// TIA Portal project "1215C_BREAKOUT_BOARD_IO-LINK_TOWERLIGHT" (V19) (continued)
REGION Network 1: ================= PORT_X1 =================
END_REGION

REGION Network 2: Reserved
END_REGION

REGION Network 3: ================= PORT_X2 =================
END_REGION

REGION Network 4: Banner Tower Light
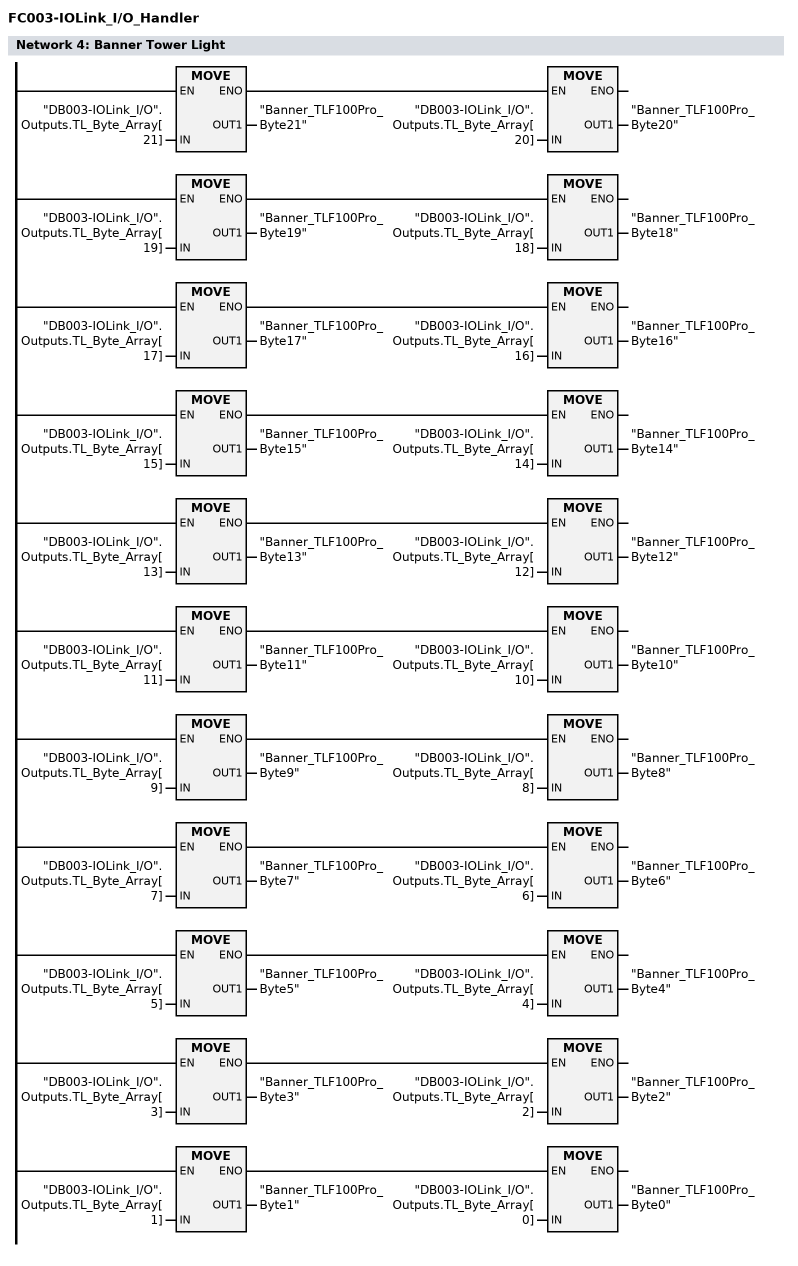
   RUNG wire#powerrail
      Move(in := "DB003-IOLink_I/O".Outputs.TL_Byte_Array[21], out1 => "Banner_TLF100Pro_Byte21")
      Move(in := "DB003-IOLink_I/O".Outputs.TL_Byte_Array[20], out1 => "Banner_TLF100Pro_Byte20")
   END_RUNG
   RUNG wire#powerrail
      Move(in := "DB003-IOLink_I/O".Outputs.TL_Byte_Array[19], out1 => "Banner_TLF100Pro_Byte19")
      Move(in := "DB003-IOLink_I/O".Outputs.TL_Byte_Array[18], out1 => "Banner_TLF100Pro_Byte18")
   END_RUNG
   RUNG wire#powerrail
      Move(in := "DB003-IOLink_I/O".Outputs.TL_Byte_Array[17], out1 => "Banner_TLF100Pro_Byte17")
      Move(in := "DB003-IOLink_I/O".Outputs.TL_Byte_Array[16], out1 => "Banner_TLF100Pro_Byte16")
   END_RUNG
   RUNG wire#powerrail
      Move(in := "DB003-IOLink_I/O".Outputs.TL_Byte_Array[15], out1 => "Banner_TLF100Pro_Byte15")
      Move(in := "DB003-IOLink_I/O".Outputs.TL_Byte_Array[14], out1 => "Banner_TLF100Pro_Byte14")
   END_RUNG
   RUNG wire#powerrail
      Move(in := "DB003-IOLink_I/O".Outputs.TL_Byte_Array[13], out1 => "Banner_TLF100Pro_Byte13")
      Move(in := "DB003-IOLink_I/O".Outputs.TL_Byte_Array[12], out1 => "Banner_TLF100Pro_Byte12")
   END_RUNG
   RUNG wire#powerrail
      Move(in := "DB003-IOLink_I/O".Outputs.TL_Byte_Array[11], out1 => "Banner_TLF100Pro_Byte11")
      Move(in := "DB003-IOLink_I/O".Outputs.TL_Byte_Array[10], out1 => "Banner_TLF100Pro_Byte10")
   END_RUNG
   RUNG wire#powerrail
      Move(in := "DB003-IOLink_I/O".Outputs.TL_Byte_Array[9], out1 => "Banner_TLF100Pro_Byte9")
      Move(in := "DB003-IOLink_I/O".Outputs.TL_Byte_Array[8], out1 => "Banner_TLF100Pro_Byte8")
   END_RUNG
   RUNG wire#powerrail
      Move(in := "DB003-IOLink_I/O".Outputs.TL_Byte_Array[7], out1 => "Banner_TLF100Pro_Byte7")
      Move(in := "DB003-IOLink_I/O".Outputs.TL_Byte_Array[6], out1 => "Banner_TLF100Pro_Byte6")
   END_RUNG
   RUNG wire#powerrail
      Move(in := "DB003-IOLink_I/O".Outputs.TL_Byte_Array[5], out1 => "Banner_TLF100Pro_Byte5")
      Move(in := "DB003-IOLink_I/O".Outputs.TL_Byte_Array[4], out1 => "Banner_TLF100Pro_Byte4")
   END_RUNG
   RUNG wire#powerrail
      Move(in := "DB003-IOLink_I/O".Outputs.TL_Byte_Array[3], out1 => "Banner_TLF100Pro_Byte3")
      Move(in := "DB003-IOLink_I/O".Outputs.TL_Byte_Array[2], out1 => "Banner_TLF100Pro_Byte2")
   END_RUNG
   RUNG wire#powerrail
      Move(in := "DB003-IOLink_I/O".Outputs.TL_Byte_Array[1], out1 => "Banner_TLF100Pro_Byte1")
      Move(in := "DB003-IOLink_I/O".Outputs.TL_Byte_Array[0], out1 => "Banner_TLF100Pro_Byte0")
   END_RUNG
   // the same network as SCL:
   "Banner_TLF100Pro_Byte21" := "DB003-IOLink_I/O".Outputs.TL_Byte_Array[21];
   "Banner_TLF100Pro_Byte20" := "DB003-IOLink_I/O".Outputs.TL_Byte_Array[20];
   "Banner_TLF100Pro_Byte19" := "DB003-IOLink_I/O".Outputs.TL_Byte_Array[19];
   "Banner_TLF100Pro_Byte18" := "DB003-IOLink_I/O".Outputs.TL_Byte_Array[18];
   "Banner_TLF100Pro_Byte17" := "DB003-IOLink_I/O".Outputs.TL_Byte_Array[17];
   "Banner_TLF100Pro_Byte16" := "DB003-IOLink_I/O".Outputs.TL_Byte_Array[16];
   "Banner_TLF100Pro_Byte15" := "DB003-IOLink_I/O".Outputs.TL_Byte_Array[15];
   "Banner_TLF100Pro_Byte14" := "DB003-IOLink_I/O".Outputs.TL_Byte_Array[14];
   "Banner_TLF100Pro_Byte13" := "DB003-IOLink_I/O".Outputs.TL_Byte_Array[13];
   "Banner_TLF100Pro_Byte12" := "DB003-IOLink_I/O".Outputs.TL_Byte_Array[12];
   "Banner_TLF100Pro_Byte11" := "DB003-IOLink_I/O".Outputs.TL_Byte_Array[11];
   "Banner_TLF100Pro_Byte10" := "DB003-IOLink_I/O".Outputs.TL_Byte_Array[10];
   "Banner_TLF100Pro_Byte9" := "DB003-IOLink_I/O".Outputs.TL_Byte_Array[9];
   "Banner_TLF100Pro_Byte8" := "DB003-IOLink_I/O".Outputs.TL_Byte_Array[8];
   "Banner_TLF100Pro_Byte7" := "DB003-IOLink_I/O".Outputs.TL_Byte_Array[7];
   "Banner_TLF100Pro_Byte6" := "DB003-IOLink_I/O".Outputs.TL_Byte_Array[6];
   "Banner_TLF100Pro_Byte5" := "DB003-IOLink_I/O".Outputs.TL_Byte_Array[5];
   "Banner_TLF100Pro_Byte4" := "DB003-IOLink_I/O".Outputs.TL_Byte_Array[4];
   "Banner_TLF100Pro_Byte3" := "DB003-IOLink_I/O".Outputs.TL_Byte_Array[3];
   "Banner_TLF100Pro_Byte2" := "DB003-IOLink_I/O".Outputs.TL_Byte_Array[2];
   "Banner_TLF100Pro_Byte1" := "DB003-IOLink_I/O".Outputs.TL_Byte_Array[1];
   "Banner_TLF100Pro_Byte0" := "DB003-IOLink_I/O".Outputs.TL_Byte_Array[0];
END_REGION

REGION Network 5: ================= PORT_X3 =================
END_REGION

REGION Network 6: Reserved
END_REGION

REGION Network 7: ================= PORT_X4 =================
END_REGION

REGION Network 8: Reserved
END_REGION
END_FUNCTION

// folder: WS01_TVET_Workstation/01-DateTime

FUNCTION "FC002-DateTime_Handler" : Void   // FC2, LAD
TITLE = Date Time Handler
{ S7_Optimized_Access := 'TRUE' }
VERSION : 0.1
// This function block is for formatting the PLC time into a format suitable for display on the HMI.
   VAR_TEMP   // added for the SCL form of the ladder/FBD networks
      _w1 : Bool;
   END_VAR
BEGIN

REGION Network 1: Read Local Date/Time
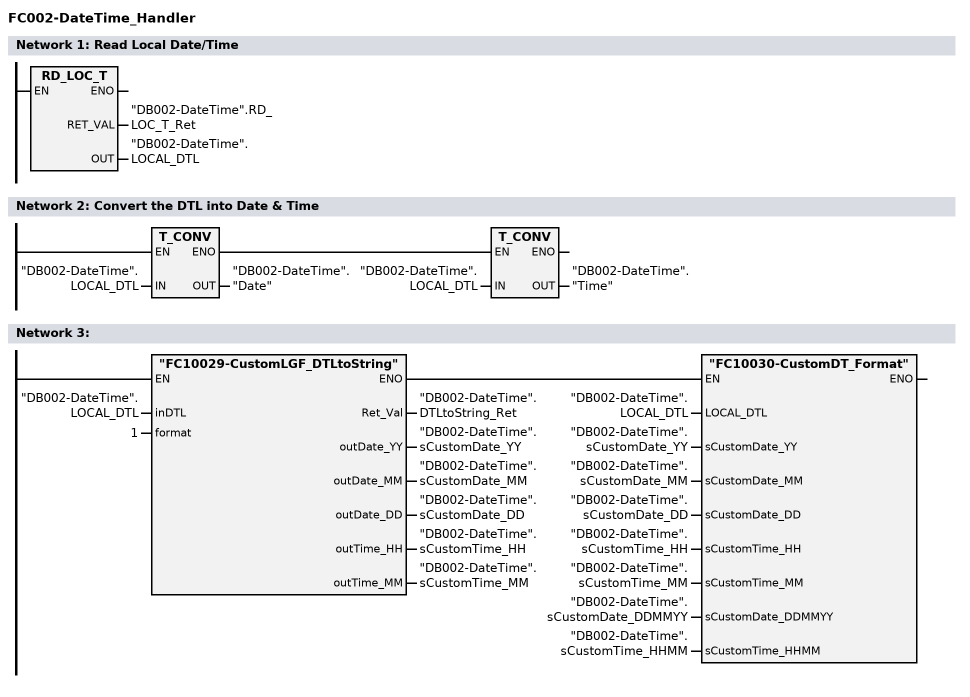
   "DB002-DateTime".RD_LOC_T_Ret := RD_LOC_T(OUT => "DB002-DateTime".LOCAL_DTL);
END_REGION

REGION Network 2: Convert the DTL into Date & Time
   // ENO of a box is taken as its EN; it also drops when the box reports an error
   "DB002-DateTime"."Date" := T_CONV(IN := "DB002-DateTime".LOCAL_DTL);
   "DB002-DateTime"."Time" := T_CONV(IN := "DB002-DateTime".LOCAL_DTL);
END_REGION

REGION Network 3
   RUNG wire#powerrail
      "FC10029-CustomLGF_DTLtoString"(inDTL := "DB002-DateTime".LOCAL_DTL, format := 1, Ret_Val => "DB002-DateTime".DTLtoString_Ret, outDate_YY => "DB002-DateTime".sCustomDate_YY, outDate_MM => "DB002-DateTime".sCustomDate_MM, outDate_DD => "DB002-DateTime".sCustomDate_DD, outTime_HH => "DB002-DateTime".sCustomTime_HH, outTime_MM => "DB002-DateTime".sCustomTime_MM)
      "FC10030-CustomDT_Format"(LOCAL_DTL := "DB002-DateTime".LOCAL_DTL, sCustomDate_YY := "DB002-DateTime".sCustomDate_YY, sCustomDate_MM := "DB002-DateTime".sCustomDate_MM, sCustomDate_DD := "DB002-DateTime".sCustomDate_DD, sCustomTime_HH := "DB002-DateTime".sCustomTime_HH, sCustomTime_MM := "DB002-DateTime".sCustomTime_MM, sCustomDate_DDMMYY := "DB002-DateTime".sCustomDate_DDMMYY, sCustomTime_HHMM := "DB002-DateTime".sCustomTime_HHMM)
   END_RUNG
   // the same network as SCL:
   "DB002-DateTime".DTLtoString_Ret := "FC10029-CustomLGF_DTLtoString"(inDTL := "DB002-DateTime".LOCAL_DTL,
                           format := 1,
                           outDate_YY => "DB002-DateTime".sCustomDate_YY,
                           outDate_MM => "DB002-DateTime".sCustomDate_MM,
                           outDate_DD => "DB002-DateTime".sCustomDate_DD,
                           outTime_HH => "DB002-DateTime".sCustomTime_HH,
                           outTime_MM => "DB002-DateTime".sCustomTime_MM,
                           ENO => #_w1);
   IF #_w1 THEN
       "FC10030-CustomDT_Format"(LOCAL_DTL := "DB002-DateTime".LOCAL_DTL,
                               sCustomDate_YY := "DB002-DateTime".sCustomDate_YY,
                               sCustomDate_MM := "DB002-DateTime".sCustomDate_MM,
                               sCustomDate_DD := "DB002-DateTime".sCustomDate_DD,
                               sCustomTime_HH := "DB002-DateTime".sCustomTime_HH,
                               sCustomTime_MM := "DB002-DateTime".sCustomTime_MM,
                               sCustomDate_DDMMYY := "DB002-DateTime".sCustomDate_DDMMYY,
                               sCustomTime_HHMM := "DB002-DateTime".sCustomTime_HHMM);
   END_IF;
END_REGION
END_FUNCTION

FUNCTION "FC10029-CustomLGF_DTLtoString" : String   // FC10029, SCL
TITLE = Custom LGF Local Date TIme to String Converter
{ S7_Optimized_Access := 'TRUE' }
VERSION : 0.1
// This function block is a modified version of the DTLtoString FC provided by Siemens in the LGF Library.
   VAR_INPUT
      inDTL : DTL;   // Date as DTL tag
      format : Bool;   // 1 = traditional, 0 = international
   END_VAR
   VAR_OUTPUT
      outDate_YY : String;   // Custom Date Output (YY)
      outDate_MM : String;   // Custom Date Output (MM)
      outDate_DD : String;   // Custom Date Output (DD)
      outTime_HH : String;   // Custom Time Output (HH)
      outTime_MM : String;   // Custom Time Output (MM)
   END_VAR
   VAR_TEMP
      tempString : String;   // -
      tempSepTime : Char;   // -
      tempPosYear : USInt;   // -
      tempPosMonth : USInt;   // -
      tempPosDay : USInt;   // -
      tempPosHour : USInt;   // -
      tempPosMinute : USInt;   // -
      tempPosSepYearMonth : USInt;   // -
      tempPosSepMonthDay : USInt;   // -
      tempPosSepHourMinute : USInt;   // -
   END_VAR
   // Ret_Val : Date as String tag
BEGIN
   //=============================================================================
   // Siemens AG
   // (c)Copyright 2017
   //-----------------------------------------------------------------------------
   // Library:       LGF (Library General Functions)
   // Tested with:   CPU1212C DC/DC/DC FW:V4.2
   // Engineering:   TIA Portal V14 Update 1
   // Restrictions:  -
   // Requirements:  PLC (S7-1200 / S7-1500)
   // Functionality: This function converts DTL into a string.  (EDITED)
   //-----------------------------------------------------------------------------
   // Change log table:
   // Version  Date        In charge / Changes applied
   // 01.00.00 15.06.2016  Siemens Industry Online Support
   //                      First released version
   // 01.00.01 02.01.2017  Siemens Industry Online Support
   //                      Upgrade: TIA Portal V14 Update 1
   // 01.00.02 17.08.2018  Siemens Industry Online Support
   //                      Upgrade: TIA V15 Update 2
   //=============================================================================


   // Initialization
   #tempString := '';
   #tempSepTime := ':';


   // Set format parameters for output string
   IF NOT #format
   THEN                                          // International ISO 8601
       #tempPosYear := 1;                          // DTL  | Y| Y| Y| Y| -| M| M| -| D| D|  | H| H| :| M| M|
       #tempPosMonth := 6;                         // -----|--|--|--|--|--|--|--|--|--|--|--|--|--|--|--|--|
       #tempPosDay := 9;                           // Pos  | 1| 2| 3| 4| 5| 6| 7| 8| 9|10|11|12|13|14|15|16|
       #tempPosHour := 12;
       #tempPosMinute := 15;
       #tempPosSepYearMonth := 5;
       #tempPosSepMonthDay := 8;
       #tempPosSepHourMinute := 14;
   ELSE                                          // Traditional (EU)
       #tempPosYear := 7;                          // DTL  | D| D| -| M| M| -| Y| Y| Y| Y|  | H| H| :| M| M|
       #tempPosMonth := 4;                         // -----|--|--|--|--|--|--|--|--|--|--|--|--|--|--|--|--|
       #tempPosDay := 1;                           // Pos  | 1| 2| 3| 4| 5| 6| 7| 8| 9|10|11|12|13|14|15|16|
       #tempPosHour := 12;
       #tempPosMinute := 15;
       #tempPosSepYearMonth := 6;
       #tempPosSepMonthDay := 3;
       #tempPosSepHourMinute := 14;
   END_IF;


   // Convert "Value" into "String" and place at the right position

   // Convert for YEAR
   VAL_STRG(FORMAT := W#16#0000,
            IN := #inDTL.YEAR,
            P := #tempPosYear,
            PREC := 0,
            SIZE := 4,
            OUT => #tempString);     // DTL YEAR --> String --> #tempPosYear

   VAL_STRG(FORMAT := W#16#0000,
            IN := #inDTL.YEAR MOD 100,
            P := 1,
            PREC := 0,
            SIZE := 2,
            OUT => #outDate_YY);        // DTL YEAR --> String --> #CustOutYear (Last 2 digits)

   // Convert for MONTH
   VAL_STRG(FORMAT := W#16#0000,
            IN := #inDTL.MONTH,
            P := #tempPosMonth,
            PREC := 0,
            SIZE := 2,
            OUT => #tempString);     // DTL MONTH --> String --> #tempPosMonth

   VAL_STRG(FORMAT := W#16#0000,
            IN := #inDTL.MONTH,
            P := 1,
            PREC := 0,
            SIZE := 2,
            OUT => #outDate_MM);        // DTL MONTH --> String --> #CustOutDate MM

   // Convert for DAY
   VAL_STRG(FORMAT := W#16#0000,
            IN := #inDTL.DAY,
            P := #tempPosDay,
            PREC := 0,
            SIZE := 2,
            OUT => #tempString);     // DTL DAY --> String --> #tempPosDay

   VAL_STRG(FORMAT := W#16#0000,
            IN := #inDTL.DAY,
            P := 1,
            PREC := 0,
            SIZE := 2,
            OUT => #outDate_DD);        // DTL DAY --> String --> #CustOutDate DDMM

   // Convert for HOUR
   VAL_STRG(FORMAT := W#16#0000,
            IN := #inDTL.HOUR,
            P := #tempPosHour,
            PREC := 0,
            SIZE := 2,
            OUT => #tempString);     // DTL HOUR --> String --> #tempPosHour

   VAL_STRG(FORMAT := W#16#0000,
            IN := #inDTL.HOUR,
            P := 1,
            PREC := 0,
            SIZE := 2,
            OUT => #outTime_HH);     // DTL HOUR --> String --> #CustOutTime HH

   // Convert for MINUTE
   VAL_STRG(FORMAT := W#16#0000,
            IN := #inDTL.MINUTE,
            P := #tempPosMinute,
            PREC := 0,
            SIZE := 2,
            OUT => #tempString);     // DTL MINUTE --> String --> #tempPosMinute

   VAL_STRG(FORMAT := W#16#0000,
            IN := #inDTL.MINUTE,
            P := 1,
            PREC := 0,
            SIZE := 2,
            OUT => #outTime_MM);        // DTL MINUTE --> String --> #CustOutTime


   // Block output
   #"FC10029-CustomLGF_DTLtoString" := #tempString;


   // Additional outputs
   #outDate_YY := #outDate_YY;
   #outDate_MM := #outDate_MM;
   #outDate_DD := #outDate_DD;
   #outTime_HH := #outTime_HH;
   #outTime_MM := #outTime_MM;
END_FUNCTION

FUNCTION "FC10030-CustomDT_Format" : Void   // FC10030, LAD
TITLE = Custom Date/Time Formats
{ S7_Optimized_Access := 'TRUE' }
VERSION : 0.1
// This function block is for formatting the local date/time display on the HMI.
   VAR_INPUT
      LOCAL_DTL : DTL;   // RAW DTL
   END_VAR
   VAR_IN_OUT
      sCustomDate_YY : String;   // Custom Year Output (YY)
      sCustomDate_MM : String;   // Custom Date Output (MM)
      sCustomDate_DD : String;   // Custom Date Output (DD)
      sCustomTime_HH : String;   // Custom Time Output (HH)
      sCustomTime_MM : String;   // Custom Time Output (MM)
      sCustomDate_DDMMYY : String;   // Custom Date (DD/MM/YY)
      sCustomTime_HHMM : String;   // Custom Date (HH:MM)
   END_VAR
   VAR_TEMP
      sTemp_String : String;   // -
   END_VAR
BEGIN

REGION Network 1: =================ADD_LEADING_ZEROS=================
END_REGION

REGION Network 2: Add leading zero to MM if less than 10
   // > If DTL.MONTH is less than 10 - replace 1st character in DD with a 0
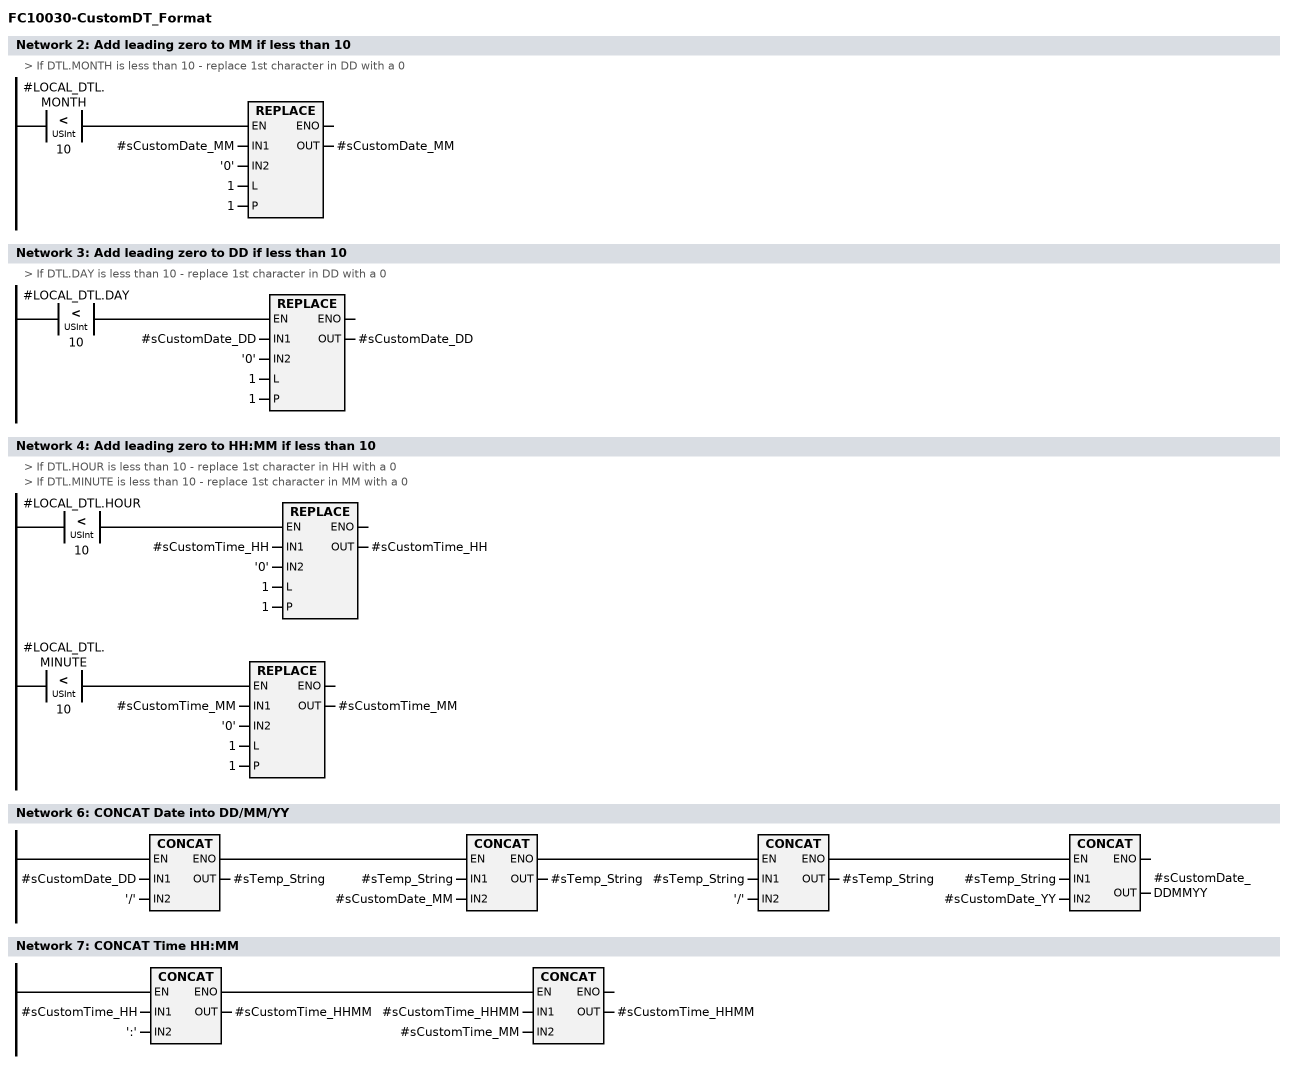
   IF #LOCAL_DTL.MONTH < 10 THEN
       #sCustomDate_MM := REPLACE(IN1 := #sCustomDate_MM, IN2 := '0', L := 1, P := 1);
   END_IF;
END_REGION

REGION Network 3: Add leading zero to DD if less than 10
   // > If DTL.DAY is less than 10 - replace 1st character in DD with a 0
   IF #LOCAL_DTL.DAY < 10 THEN
       #sCustomDate_DD := REPLACE(IN1 := #sCustomDate_DD, IN2 := '0', L := 1, P := 1);
   END_IF;
END_REGION

REGION Network 4: Add leading zero to HH:MM if less than 10
   // > If DTL.HOUR is less than 10 - replace 1st character in HH with a 0
   // > If DTL.MINUTE is less than 10 - replace 1st character in MM with a 0
   IF #LOCAL_DTL.HOUR < 10 THEN
       #sCustomTime_HH := REPLACE(IN1 := #sCustomTime_HH, IN2 := '0', L := 1, P := 1);
   END_IF;
   IF #LOCAL_DTL.MINUTE < 10 THEN
       #sCustomTime_MM := REPLACE(IN1 := #sCustomTime_MM, IN2 := '0', L := 1, P := 1);
   END_IF;
END_REGION

REGION Network 5: =================CONCAT_INTO_FORMAT=================
END_REGION

REGION Network 6: CONCAT Date into DD/MM/YY
   #sTemp_String := CONCAT(IN1 := #sCustomDate_DD, IN2 := '/');
   #sTemp_String := CONCAT(IN1 := #sTemp_String, IN2 := #sCustomDate_MM);
   #sTemp_String := CONCAT(IN1 := #sTemp_String, IN2 := '/');
   #sCustomDate_DDMMYY := CONCAT(IN1 := #sTemp_String, IN2 := #sCustomDate_YY);
END_REGION

REGION Network 7: CONCAT Time HH:MM
   #sCustomTime_HHMM := CONCAT(IN1 := #sCustomTime_HH, IN2 := ':');
   #sCustomTime_HHMM := CONCAT(IN1 := #sCustomTime_HHMM, IN2 := #sCustomTime_MM);
END_REGION
END_FUNCTION

// folder: WS01_TVET_Workstation/02-IOLink_Control

FUNCTION "FC004-TowerLight_Handler" : Void   // FC4, LAD
TITLE = IOLink Tower Light Control
{ S7_Optimized_Access := 'TRUE' }
VERSION : 0.1
// This function block is for switching the tower light segments ON or OFF, which are configured via the HMI panel.
   VAR_OUTPUT
      TL_Byte_Array : Array[0..21] of Byte;   // Tower Light Byte Array
   END_VAR
BEGIN

REGION Network 1: ================= SEGMENT_ONE =================
END_REGION

REGION Network 2: OFF
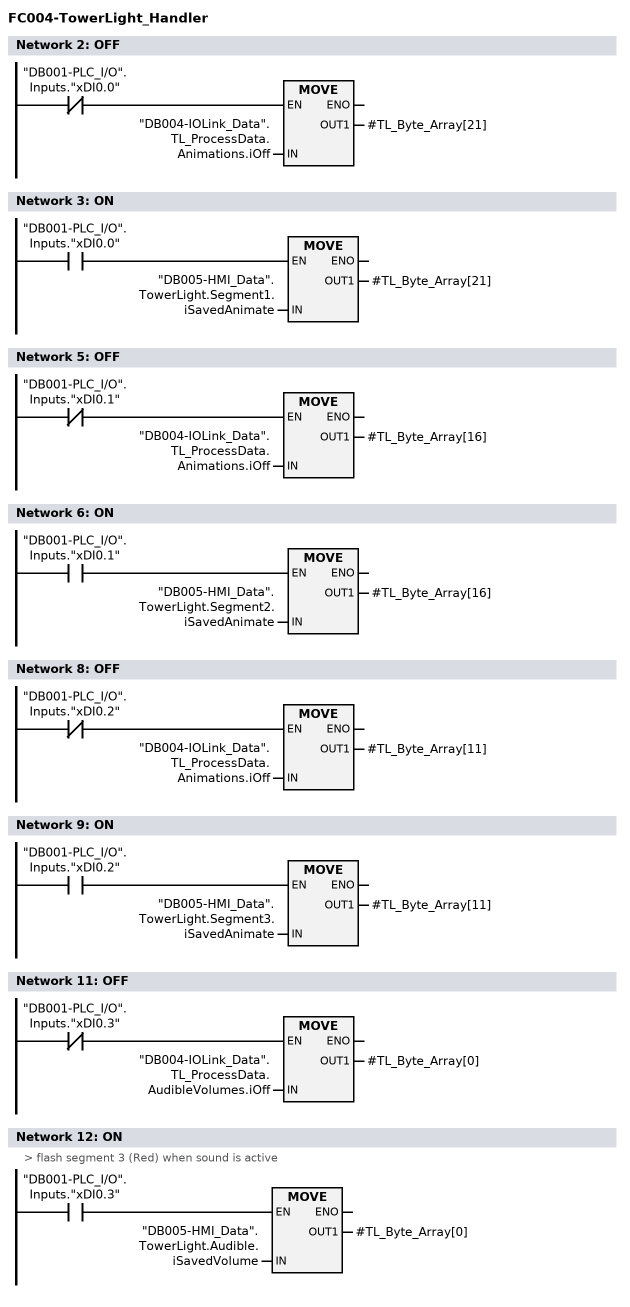
   RUNG wire#powerrail
      I_Contact( "DB001-PLC_I/O".Inputs."xDI0.0" )
      Move(in := "DB004-IOLink_Data".TL_ProcessData.Animations.iOff, out1 => #TL_Byte_Array[21])
   END_RUNG
   // the same network as SCL:
   IF NOT "DB001-PLC_I/O".Inputs."xDI0.0" THEN
       #TL_Byte_Array[21] := "DB004-IOLink_Data".TL_ProcessData.Animations.iOff;
   END_IF;
END_REGION

REGION Network 3: ON
   RUNG wire#powerrail
      Contact( "DB001-PLC_I/O".Inputs."xDI0.0" )
      Move(in := "DB005-HMI_Data".TowerLight.Segment1.iSavedAnimate, out1 => #TL_Byte_Array[21])
   END_RUNG
   // the same network as SCL:
   IF "DB001-PLC_I/O".Inputs."xDI0.0" THEN
       #TL_Byte_Array[21] := "DB005-HMI_Data".TowerLight.Segment1.iSavedAnimate;
   END_IF;
END_REGION

REGION Network 4: ================= SEGMENT_TWO =================
END_REGION

REGION Network 5: OFF
   RUNG wire#powerrail
      I_Contact( "DB001-PLC_I/O".Inputs."xDI0.1" )
      Move(in := "DB004-IOLink_Data".TL_ProcessData.Animations.iOff, out1 => #TL_Byte_Array[16])
   END_RUNG
   // the same network as SCL:
   IF NOT "DB001-PLC_I/O".Inputs."xDI0.1" THEN
       #TL_Byte_Array[16] := "DB004-IOLink_Data".TL_ProcessData.Animations.iOff;
   END_IF;
END_REGION

REGION Network 6: ON
   RUNG wire#powerrail
      Contact( "DB001-PLC_I/O".Inputs."xDI0.1" )
      Move(in := "DB005-HMI_Data".TowerLight.Segment2.iSavedAnimate, out1 => #TL_Byte_Array[16])
   END_RUNG
   // the same network as SCL:
   IF "DB001-PLC_I/O".Inputs."xDI0.1" THEN
       #TL_Byte_Array[16] := "DB005-HMI_Data".TowerLight.Segment2.iSavedAnimate;
   END_IF;
END_REGION

REGION Network 7: ================= SEGMENT_THREE =================
END_REGION

REGION Network 8: OFF
   RUNG wire#powerrail
      I_Contact( "DB001-PLC_I/O".Inputs."xDI0.2" )
      Move(in := "DB004-IOLink_Data".TL_ProcessData.Animations.iOff, out1 => #TL_Byte_Array[11])
   END_RUNG
   // the same network as SCL:
   IF NOT "DB001-PLC_I/O".Inputs."xDI0.2" THEN
       #TL_Byte_Array[11] := "DB004-IOLink_Data".TL_ProcessData.Animations.iOff;
   END_IF;
END_REGION

REGION Network 9: ON
   RUNG wire#powerrail
      Contact( "DB001-PLC_I/O".Inputs."xDI0.2" )
      Move(in := "DB005-HMI_Data".TowerLight.Segment3.iSavedAnimate, out1 => #TL_Byte_Array[11])
   END_RUNG
   // the same network as SCL:
   IF "DB001-PLC_I/O".Inputs."xDI0.2" THEN
       #TL_Byte_Array[11] := "DB005-HMI_Data".TowerLight.Segment3.iSavedAnimate;
   END_IF;
END_REGION

REGION Network 10: ================= AUDIBLE =================
END_REGION

REGION Network 11: OFF
   RUNG wire#powerrail
      I_Contact( "DB001-PLC_I/O".Inputs."xDI0.3" )
      Move(in := "DB004-IOLink_Data".TL_ProcessData.AudibleVolumes.iOff, out1 => #TL_Byte_Array[0])
   END_RUNG
   // the same network as SCL:
   IF NOT "DB001-PLC_I/O".Inputs."xDI0.3" THEN
       #TL_Byte_Array[0] := "DB004-IOLink_Data".TL_ProcessData.AudibleVolumes.iOff;
   END_IF;
END_REGION

REGION Network 12: ON
   // > flash segment 3 (Red) when sound is active
   RUNG wire#powerrail
      Contact( "DB001-PLC_I/O".Inputs."xDI0.3" )
      Move(in := "DB005-HMI_Data".TowerLight.Audible.iSavedVolume, out1 => #TL_Byte_Array[0])
   END_RUNG
   // the same network as SCL:
   IF "DB001-PLC_I/O".Inputs."xDI0.3" THEN
       #TL_Byte_Array[0] := "DB005-HMI_Data".TowerLight.Audible.iSavedVolume;
   END_IF;
END_REGION
END_FUNCTION

// folder: WS01_TVET_Workstation/03-HMI_Control

FUNCTION "FC005-HMI_Handler" : Void   // FC5, LAD
TITLE = HMI Data Handler
{ S7_Optimized_Access := 'TRUE' }
VERSION : 0.1
// This function block is for interfacing HMI data to a Global DB (DB005-HMI_Data).
   VAR_OUTPUT
      TL_Byte_Array : Array[0..21] of Byte;   // Tower Light Byte Array
   END_VAR
   VAR_TEMP
      Seg1 : Struct
         iTempAnimation : Int;
         iTempSpeed : Int;
         iTempColour1 : Int;
         iTempColour2 : Int;
         "iTempClrWidth%" : Int;
      END_STRUCT;
      Seg2 : Struct
         iTempAnimation : Int;
         iTempSpeed : Int;
         iTempColour1 : Int;
         iTempColour2 : Int;
         "iTempClrWidth%" : Int;
      END_STRUCT;
      Seg3 : Struct
         iTempAnimation : Int;
         iTempSpeed : Int;
         iTempColour1 : Int;
         iTempColour2 : Int;
         "iTempClrWidth%" : Int;
      END_STRUCT;
      Audible : Struct
         iTempType : Int;
         iTempVolume : Int;
      END_STRUCT;
   END_VAR
BEGIN

REGION Network 1: ================= SEGMENT_ONE =================
END_REGION

REGION Network 2: While making selections
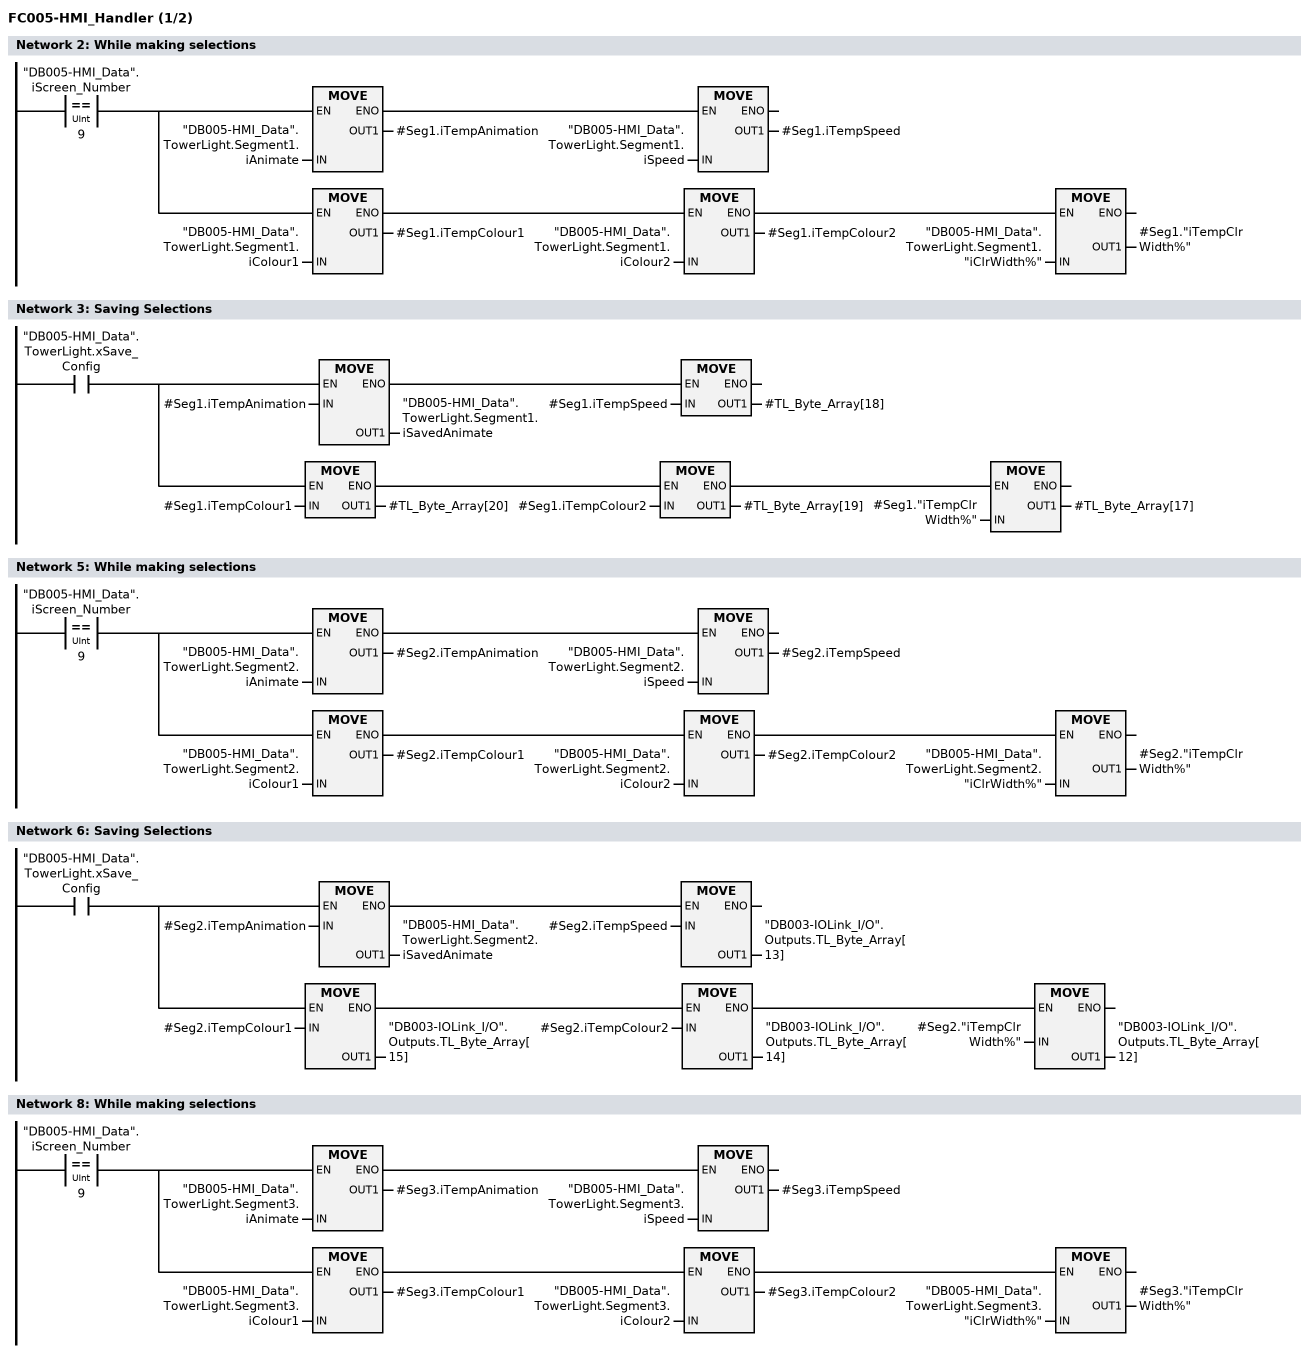
   RUNG wire#powerrail
      { S7_Templates := "SrcType := UInt" } EQ_Contact(in1 := "DB005-HMI_Data".iScreen_Number, in2 := 9)
      wire#w1
      Move(in := "DB005-HMI_Data".TowerLight.Segment1.iAnimate, out1 => #Seg1.iTempAnimation)
      Move(in := "DB005-HMI_Data".TowerLight.Segment1.iSpeed, out1 => #Seg1.iTempSpeed)
   END_RUNG
   RUNG wire#w1
      Move(in := "DB005-HMI_Data".TowerLight.Segment1.iColour1, out1 => #Seg1.iTempColour1)
      Move(in := "DB005-HMI_Data".TowerLight.Segment1.iColour2, out1 => #Seg1.iTempColour2)
      Move(in := "DB005-HMI_Data".TowerLight.Segment1."iClrWidth%", out1 => #Seg1."iTempClrWidth%")
   END_RUNG
   // the same network as SCL:
   IF "DB005-HMI_Data".iScreen_Number = 9 THEN
       #Seg1.iTempAnimation := "DB005-HMI_Data".TowerLight.Segment1.iAnimate;
       #Seg1.iTempSpeed := "DB005-HMI_Data".TowerLight.Segment1.iSpeed;
       #Seg1.iTempColour1 := "DB005-HMI_Data".TowerLight.Segment1.iColour1;
       #Seg1.iTempColour2 := "DB005-HMI_Data".TowerLight.Segment1.iColour2;
       #Seg1."iTempClrWidth%" := "DB005-HMI_Data".TowerLight.Segment1."iClrWidth%";
   END_IF;
END_REGION

REGION Network 3: Saving Selections
   RUNG wire#powerrail
      Contact( "DB005-HMI_Data".TowerLight.xSave_Config )
      wire#w1
      Move(in := #Seg1.iTempAnimation, out1 => "DB005-HMI_Data".TowerLight.Segment1.iSavedAnimate)
      Move(in := #Seg1.iTempSpeed, out1 => #TL_Byte_Array[18])
   END_RUNG
   RUNG wire#w1
      Move(in := #Seg1.iTempColour1, out1 => #TL_Byte_Array[20])
      Move(in := #Seg1.iTempColour2, out1 => #TL_Byte_Array[19])
      Move(in := #Seg1."iTempClrWidth%", out1 => #TL_Byte_Array[17])
   END_RUNG
   // the same network as SCL:
   IF "DB005-HMI_Data".TowerLight.xSave_Config THEN
       "DB005-HMI_Data".TowerLight.Segment1.iSavedAnimate := #Seg1.iTempAnimation;
       #TL_Byte_Array[18] := #Seg1.iTempSpeed;
       #TL_Byte_Array[20] := #Seg1.iTempColour1;
       #TL_Byte_Array[19] := #Seg1.iTempColour2;
       #TL_Byte_Array[17] := #Seg1."iTempClrWidth%";
   END_IF;
END_REGION

REGION Network 4: ================= SEGMENT_TWO =================
END_REGION

REGION Network 5: While making selections
   RUNG wire#powerrail
      { S7_Templates := "SrcType := UInt" } EQ_Contact(in1 := "DB005-HMI_Data".iScreen_Number, in2 := 9)
      wire#w1
      Move(in := "DB005-HMI_Data".TowerLight.Segment2.iAnimate, out1 => #Seg2.iTempAnimation)
      Move(in := "DB005-HMI_Data".TowerLight.Segment2.iSpeed, out1 => #Seg2.iTempSpeed)
   END_RUNG
   RUNG wire#w1
      Move(in := "DB005-HMI_Data".TowerLight.Segment2.iColour1, out1 => #Seg2.iTempColour1)
      Move(in := "DB005-HMI_Data".TowerLight.Segment2.iColour2, out1 => #Seg2.iTempColour2)
      Move(in := "DB005-HMI_Data".TowerLight.Segment2."iClrWidth%", out1 => #Seg2."iTempClrWidth%")
   END_RUNG
   // the same network as SCL:
   IF "DB005-HMI_Data".iScreen_Number = 9 THEN
       #Seg2.iTempAnimation := "DB005-HMI_Data".TowerLight.Segment2.iAnimate;
       #Seg2.iTempSpeed := "DB005-HMI_Data".TowerLight.Segment2.iSpeed;
       #Seg2.iTempColour1 := "DB005-HMI_Data".TowerLight.Segment2.iColour1;
       #Seg2.iTempColour2 := "DB005-HMI_Data".TowerLight.Segment2.iColour2;
       #Seg2."iTempClrWidth%" := "DB005-HMI_Data".TowerLight.Segment2."iClrWidth%";
   END_IF;
END_REGION
